REGION Network 2: Orden de marcha desde Panel MC002 - Compresor de Alta ABC3
   RUNG wire#powerrail
      Contact( "PanelCmpAlta".MarchaPanelMC002 )
      I_Contact( "PanelCmpAlta".MantMC002 )
      Coil( "DB-CompAltaDatos".PanMchCmp2 )
   END_RUNG
   // the same network as SCL:
   "DB-CompAltaDatos".PanMchCmp2 := "PanelCmpAlta".MarchaPanelMC002 AND NOT "PanelCmpAlta".MantMC002;
END_REGION

REGION Network 3: Orden de marcha desde Panel MC003 - Compresor de Alta BELLIS
   RUNG wire#powerrail
      Contact( "PanelCmpAlta".MarchaPanelMC003 )
      I_Contact( "PanelCmpAlta".MantMC003 )
      Coil( "DB-CompAltaDatos".PanMchCmp3 )
   END_RUNG
   // the same network as SCL:
   "DB-CompAltaDatos".PanMchCmp3 := "PanelCmpAlta".MarchaPanelMC003 AND NOT "PanelCmpAlta".MantMC003;
END_REGION

REGION Network 4: Orden de marcha desde Panel MC004 - Compresor de Alta ABC4
   RUNG wire#powerrail
      Contact( "PanelCmpAlta".MarchaPanelMC004 )
      I_Contact( "PanelCmpAlta".MantMC004 )
      Coil( "DB-CompAltaDatos".PanMchCmp4 )
   END_RUNG
   // the same network as SCL:
   "DB-CompAltaDatos".PanMchCmp4 := "PanelCmpAlta".MarchaPanelMC004 AND NOT "PanelCmpAlta".MantMC004;
END_REGION

REGION Network 5: Orden de marcha desde Panel MC005 - Compresor de Alta ABC5
   RUNG wire#powerrail
      Contact( "PanelCmpAlta".MarchaPanelMC005 )
      I_Contact( "PanelCmpAlta".MantMC005 )
      Coil( "DB-CompAltaDatos".PanMchCmp5 )
   END_RUNG
   // the same network as SCL:
   "DB-CompAltaDatos".PanMchCmp5 := "PanelCmpAlta".MarchaPanelMC005 AND NOT "PanelCmpAlta".MantMC005;
END_REGION

REGION Network 6: Orden de marcha desde Panel MC005 - Compresor de Alta ABC5
   RUNG wire#powerrail
      Contact( "PanelCmpAlta".MarchaPanelMC006 )
      I_Contact( "PanelCmpAlta".MantMC006 )
      Coil( "DB-CompAltaDatos".PanMchCmp6 )
   END_RUNG
   // the same network as SCL:
   "DB-CompAltaDatos".PanMchCmp6 := "PanelCmpAlta".MarchaPanelMC006 AND NOT "PanelCmpAlta".MantMC006;
END_REGION

REGION Network 7: Salida de mantenimiento compresor 1 / Mantenimiento MC001 - Compresor de Alta ABC2
   RUNG wire#powerrail
      Contact( "PanelCmpAlta".MantMC001 )
      Not()
      Coil( "MC001_MANT" )
   END_RUNG
   // the same network as SCL:
   "MC001_MANT" := NOT "PanelCmpAlta".MantMC001;
END_REGION

REGION Network 8: Salida de mantenimiento compresor 2 / Mantenimiento MC002 - Compresor de Alta ABC3
   RUNG wire#powerrail
      Contact( "PanelCmpAlta".MantMC002 )
      Not()
      Coil( "MC002_MANT" )
   END_RUNG
   // the same network as SCL:
   "MC002_MANT" := NOT "PanelCmpAlta".MantMC002;
END_REGION

REGION Network 9: Salida de mantenimiento compresor 3 / Mantenimiento MC003 - Compresor de Alta BELLIS
   RUNG wire#powerrail
      Contact( "PanelCmpAlta".MantMC003 )
      Not()
      Coil( "MC003_MANT" )
   END_RUNG
   // the same network as SCL:
   "MC003_MANT" := NOT "PanelCmpAlta".MantMC003;
END_REGION

REGION Network 10: Salida de mantenimiento compresor 4 / Mantenimiento MC004 - Compresor de Alta ABC4
   RUNG wire#powerrail
      Contact( "PanelCmpAlta".MantMC004 )
      Not()
      Coil( "MC004_MANT" )
   END_RUNG
   // the same network as SCL:
   "MC004_MANT" := NOT "PanelCmpAlta".MantMC004;
END_REGION

REGION Network 11: Salida de mantenimiento compresor 5 / Mantenimiento MC005 - Compresor de Alta ABC5
   RUNG wire#powerrail
      Contact( "PanelCmpAlta".MantMC005 )
      Not()
      Coil( "MC005_MANT" )
   END_RUNG
   // the same network as SCL:
   "MC005_MANT" := NOT "PanelCmpAlta".MantMC005;
END_REGION

REGION Network 12: Salida de mantenimiento compresor 6 / Mantenimiento MC005 - Compresor de Alta ABC5
   RUNG wire#powerrail
      Contact( "PanelCmpAlta".MantMC006 )
      Not()
      Coil( "MC006_MANT" )
   END_RUNG
   // the same network as SCL:
   "MC006_MANT" := NOT "PanelCmpAlta".MantMC006;
END_REGION

REGION Network 13: Aparentemente obsoleto
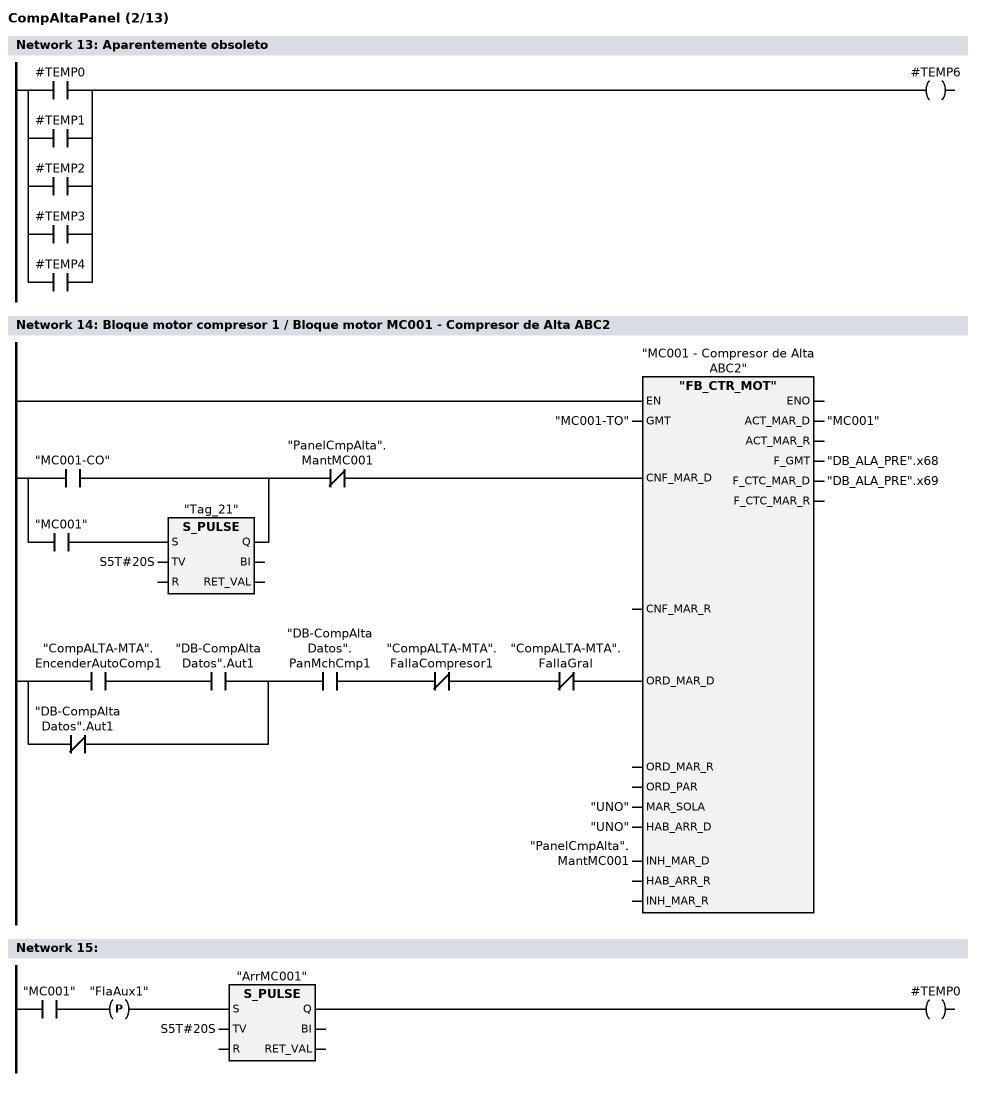
   RUNG wire#powerrail
      Contact( #TEMP0 )
      wire#w1
      Coil( #TEMP6 )
   END_RUNG
   RUNG wire#powerrail
      Contact( #TEMP1 )
   END_RUNG wire#w1
   RUNG wire#powerrail
      Contact( #TEMP2 )
   END_RUNG wire#w1
   RUNG wire#powerrail
      Contact( #TEMP3 )
   END_RUNG wire#w1
   RUNG wire#powerrail
      Contact( #TEMP4 )
   END_RUNG wire#w1
   // the same network as SCL:
   #TEMP6 := #TEMP0 OR #TEMP1 OR #TEMP2 OR #TEMP3 OR #TEMP4;
END_REGION

REGION Network 14: Bloque motor compresor 1 / Bloque motor MC001 - Compresor de Alta ABC2
   RUNG wire#powerrail
      "MC001 - Compresor de Alta ABC2"(CNF_MAR_D := wire#w2, ORD_MAR_D := wire#w4, GMT := "MC001-TO", CNF_MAR_R :=, ORD_MAR_R :=, ORD_PAR :=, MAR_SOLA := "UNO", HAB_ARR_D := "UNO", INH_MAR_D := "PanelCmpAlta".MantMC001, HAB_ARR_R :=, INH_MAR_R :=, ACT_MAR_D => "MC001", ACT_MAR_R =>, F_GMT => "DB_ALA_PRE".x68, F_CTC_MAR_D => "DB_ALA_PRE".x69, F_CTC_MAR_R =>)
   END_RUNG
   RUNG wire#powerrail
      Contact( "MC001-CO" )
      wire#w1
      I_Contact( "PanelCmpAlta".MantMC001 )
   END_RUNG wire#w2
   RUNG wire#powerrail
      Contact( "MC001" )
      S_PULSE(T_NO := "Tag_21", TV := S5T#20S, R :=, BI =>, RET_VAL =>)
   END_RUNG wire#w1
   RUNG wire#powerrail
      Contact( "CompALTA-MTA".EncenderAutoComp1 )
      Contact( "DB-CompAltaDatos".Aut1 )
      wire#w3
      Contact( "DB-CompAltaDatos".PanMchCmp1 )
      I_Contact( "CompALTA-MTA".FallaCompresor1 )
      I_Contact( "CompALTA-MTA".FallaGral )
   END_RUNG wire#w4
   RUNG wire#powerrail
      I_Contact( "DB-CompAltaDatos".Aut1 )
   END_RUNG wire#w3
   // the same network as SCL:
   #_s5time1 := S_PULSE(T_NO := "Tag_21", S := "MC001", TV := S5T#20S, Q => #_w1);
   "MC001 - Compresor de Alta ABC2"(GMT := "MC001-TO",   // "FB_CTR_MOT"
                           CNF_MAR_D := ("MC001-CO" OR #_w1) AND NOT "PanelCmpAlta".MantMC001,
                           ORD_MAR_D := (("CompALTA-MTA".EncenderAutoComp1 AND "DB-CompAltaDatos".Aut1) OR NOT "DB-CompAltaDatos".Aut1) AND "DB-CompAltaDatos".PanMchCmp1 AND NOT "CompALTA-MTA".FallaCompresor1 AND NOT "CompALTA-MTA".FallaGral,
                           MAR_SOLA := "UNO",
                           HAB_ARR_D := "UNO",
                           INH_MAR_D := "PanelCmpAlta".MantMC001,
                           ACT_MAR_D => "MC001",
                           F_GMT => "DB_ALA_PRE".x68,
                           F_CTC_MAR_D => "DB_ALA_PRE".x69);
END_REGION

REGION Network 15
   RUNG wire#powerrail
      Contact( "MC001" )
      P_Trig( "FlaAux1" )
      S_PULSE(T_NO := "ArrMC001", TV := S5T#20S, R :=, BI =>, RET_VAL =>)
      Coil( #TEMP0 )
   END_RUNG
   // the same network as SCL:
   #_w1 := "MC001" AND NOT "FlaAux1";   // rising edge
   "FlaAux1" := "MC001";
   #_s5time1 := S_PULSE(T_NO := "ArrMC001", S := #_w1, TV := S5T#20S, Q => #_w2);
   #TEMP0 := #_w2;
END_REGION

REGION Network 16: Bloque motor compresor 2 / Bloque motor MC002 - Compresor de Alta ABC3
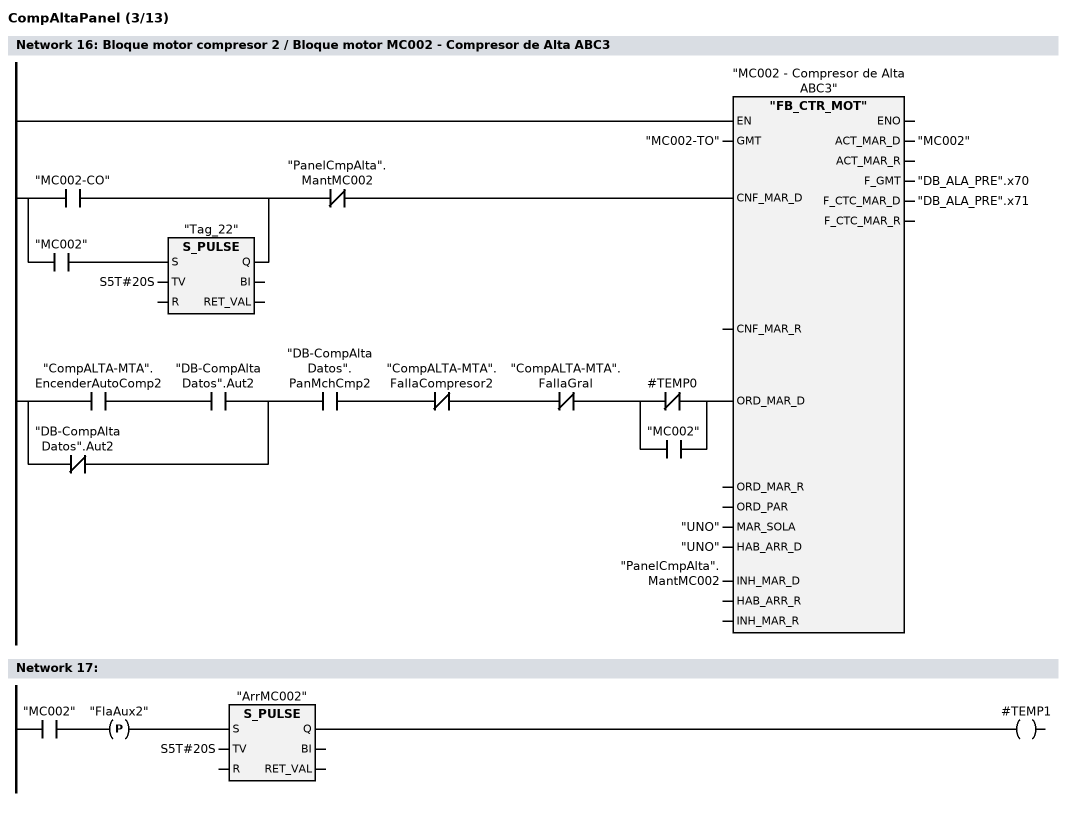
   RUNG wire#powerrail
      "MC002 - Compresor de Alta ABC3"(CNF_MAR_D := wire#w2, ORD_MAR_D := wire#w5, GMT := "MC002-TO", CNF_MAR_R :=, ORD_MAR_R :=, ORD_PAR :=, MAR_SOLA := "UNO", HAB_ARR_D := "UNO", INH_MAR_D := "PanelCmpAlta".MantMC002, HAB_ARR_R :=, INH_MAR_R :=, ACT_MAR_D => "MC002", ACT_MAR_R =>, F_GMT => "DB_ALA_PRE".x70, F_CTC_MAR_D => "DB_ALA_PRE".x71, F_CTC_MAR_R =>)
   END_RUNG
   RUNG wire#powerrail
      Contact( "MC002-CO" )
      wire#w1
      I_Contact( "PanelCmpAlta".MantMC002 )
   END_RUNG wire#w2
   RUNG wire#powerrail
      Contact( "MC002" )
      S_PULSE(T_NO := "Tag_22", TV := S5T#20S, R :=, BI =>, RET_VAL =>)
   END_RUNG wire#w1
   RUNG wire#powerrail
      Contact( "CompALTA-MTA".EncenderAutoComp2 )
      Contact( "DB-CompAltaDatos".Aut2 )
      wire#w3
      Contact( "DB-CompAltaDatos".PanMchCmp2 )
      I_Contact( "CompALTA-MTA".FallaCompresor2 )
      I_Contact( "CompALTA-MTA".FallaGral )
      wire#w4
      I_Contact( #TEMP0 )
   END_RUNG wire#w5
   RUNG wire#powerrail
      I_Contact( "DB-CompAltaDatos".Aut2 )
   END_RUNG wire#w3
   RUNG wire#w4
      Contact( "MC002" )
   END_RUNG wire#w5
   // the same network as SCL:
   #_s5time1 := S_PULSE(T_NO := "Tag_22", S := "MC002", TV := S5T#20S, Q => #_w1);
   "MC002 - Compresor de Alta ABC3"(GMT := "MC002-TO",   // "FB_CTR_MOT"
                           CNF_MAR_D := ("MC002-CO" OR #_w1) AND NOT "PanelCmpAlta".MantMC002,
                           ORD_MAR_D := (("CompALTA-MTA".EncenderAutoComp2 AND "DB-CompAltaDatos".Aut2) OR NOT "DB-CompAltaDatos".Aut2) AND "DB-CompAltaDatos".PanMchCmp2 AND NOT "CompALTA-MTA".FallaCompresor2 AND NOT "CompALTA-MTA".FallaGral AND (NOT #TEMP0 OR "MC002"),
                           MAR_SOLA := "UNO",
                           HAB_ARR_D := "UNO",
                           INH_MAR_D := "PanelCmpAlta".MantMC002,
                           ACT_MAR_D => "MC002",
                           F_GMT => "DB_ALA_PRE".x70,
                           F_CTC_MAR_D => "DB_ALA_PRE".x71);
END_REGION

REGION Network 17
   RUNG wire#powerrail
      Contact( "MC002" )
      P_Trig( "FlaAux2" )
      S_PULSE(T_NO := "ArrMC002", TV := S5T#20S, R :=, BI =>, RET_VAL =>)
      Coil( #TEMP1 )
   END_RUNG
   // the same network as SCL:
   #_w1 := "MC002" AND NOT "FlaAux2";   // rising edge
   "FlaAux2" := "MC002";
   #_s5time1 := S_PULSE(T_NO := "ArrMC002", S := #_w1, TV := S5T#20S, Q => #_w2);
   #TEMP1 := #_w2;
END_REGION

REGION Network 18: Bloque motor compresor 3 / Bloque motor MC003 - Compresor de Alta BELLIS
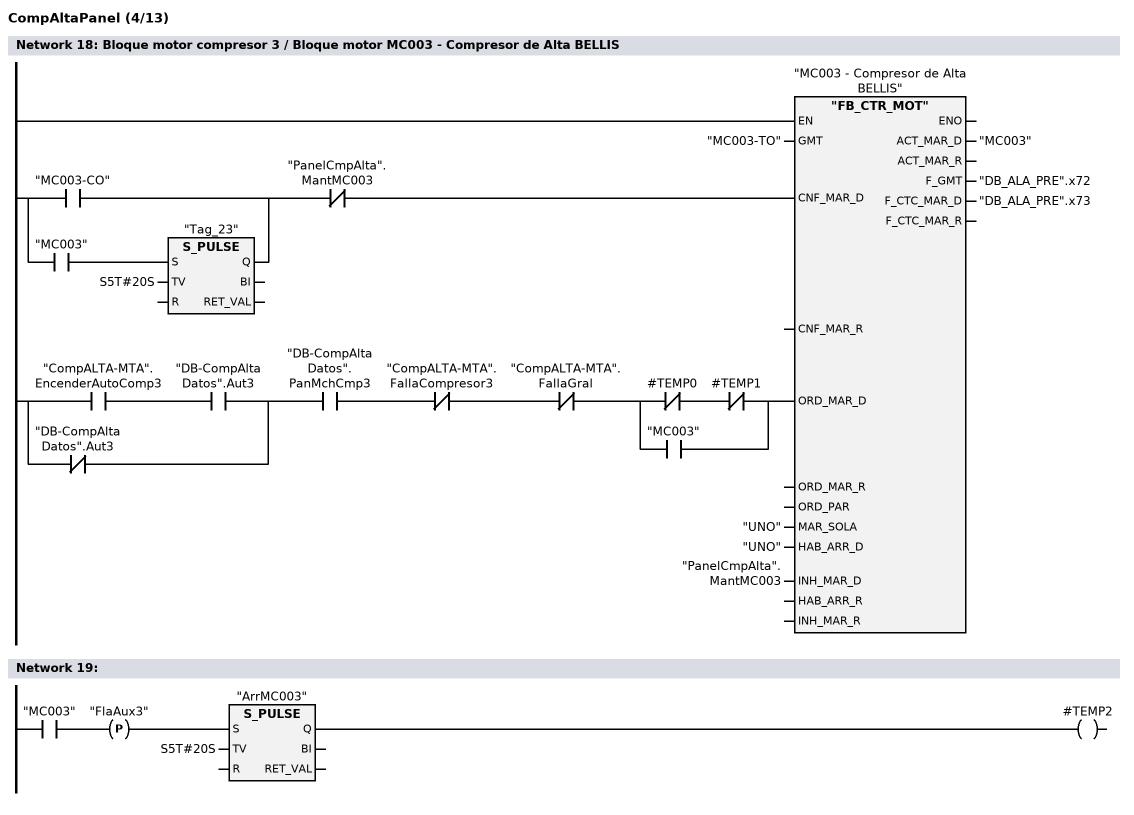
   RUNG wire#powerrail
      "MC003 - Compresor de Alta BELLIS"(CNF_MAR_D := wire#w2, ORD_MAR_D := wire#w5, GMT := "MC003-TO", CNF_MAR_R :=, ORD_MAR_R :=, ORD_PAR :=, MAR_SOLA := "UNO", HAB_ARR_D := "UNO", INH_MAR_D := "PanelCmpAlta".MantMC003, HAB_ARR_R :=, INH_MAR_R :=, ACT_MAR_D => "MC003", ACT_MAR_R =>, F_GMT => "DB_ALA_PRE".x72, F_CTC_MAR_D => "DB_ALA_PRE".x73, F_CTC_MAR_R =>)
   END_RUNG
   RUNG wire#powerrail
      Contact( "MC003-CO" )
      wire#w1
      I_Contact( "PanelCmpAlta".MantMC003 )
   END_RUNG wire#w2
   RUNG wire#powerrail
      Contact( "MC003" )
      S_PULSE(T_NO := "Tag_23", TV := S5T#20S, R :=, BI =>, RET_VAL =>)
   END_RUNG wire#w1
   RUNG wire#powerrail
      Contact( "CompALTA-MTA".EncenderAutoComp3 )
      Contact( "DB-CompAltaDatos".Aut3 )
      wire#w3
      Contact( "DB-CompAltaDatos".PanMchCmp3 )
      I_Contact( "CompALTA-MTA".FallaCompresor3 )
      I_Contact( "CompALTA-MTA".FallaGral )
      wire#w4
      I_Contact( #TEMP0 )
      I_Contact( #TEMP1 )
   END_RUNG wire#w5
   RUNG wire#powerrail
      I_Contact( "DB-CompAltaDatos".Aut3 )
   END_RUNG wire#w3
   RUNG wire#w4
      Contact( "MC003" )
   END_RUNG wire#w5
   // the same network as SCL:
   #_s5time1 := S_PULSE(T_NO := "Tag_23", S := "MC003", TV := S5T#20S, Q => #_w1);
   "MC003 - Compresor de Alta BELLIS"(GMT := "MC003-TO",   // "FB_CTR_MOT"
                           CNF_MAR_D := ("MC003-CO" OR #_w1) AND NOT "PanelCmpAlta".MantMC003,
                           ORD_MAR_D := (("CompALTA-MTA".EncenderAutoComp3 AND "DB-CompAltaDatos".Aut3) OR NOT "DB-CompAltaDatos".Aut3) AND "DB-CompAltaDatos".PanMchCmp3 AND NOT "CompALTA-MTA".FallaCompresor3 AND NOT "CompALTA-MTA".FallaGral AND ((NOT #TEMP0 AND NOT #TEMP1) OR "MC003"),
                           MAR_SOLA := "UNO",
                           HAB_ARR_D := "UNO",
                           INH_MAR_D := "PanelCmpAlta".MantMC003,
                           ACT_MAR_D => "MC003",
                           F_GMT => "DB_ALA_PRE".x72,
                           F_CTC_MAR_D => "DB_ALA_PRE".x73);
END_REGION

REGION Network 19
   RUNG wire#powerrail
      Contact( "MC003" )
      P_Trig( "FlaAux3" )
      S_PULSE(T_NO := "ArrMC003", TV := S5T#20S, R :=, BI =>, RET_VAL =>)
      Coil( #TEMP2 )
   END_RUNG
   // the same network as SCL:
   #_w1 := "MC003" AND NOT "FlaAux3";   // rising edge
   "FlaAux3" := "MC003";
   #_s5time1 := S_PULSE(T_NO := "ArrMC003", S := #_w1, TV := S5T#20S, Q => #_w2);
   #TEMP2 := #_w2;
END_REGION

REGION Network 20: Bloque motor compresor 4 / Bloque motor MC004 - Compresor de Alta ABC4
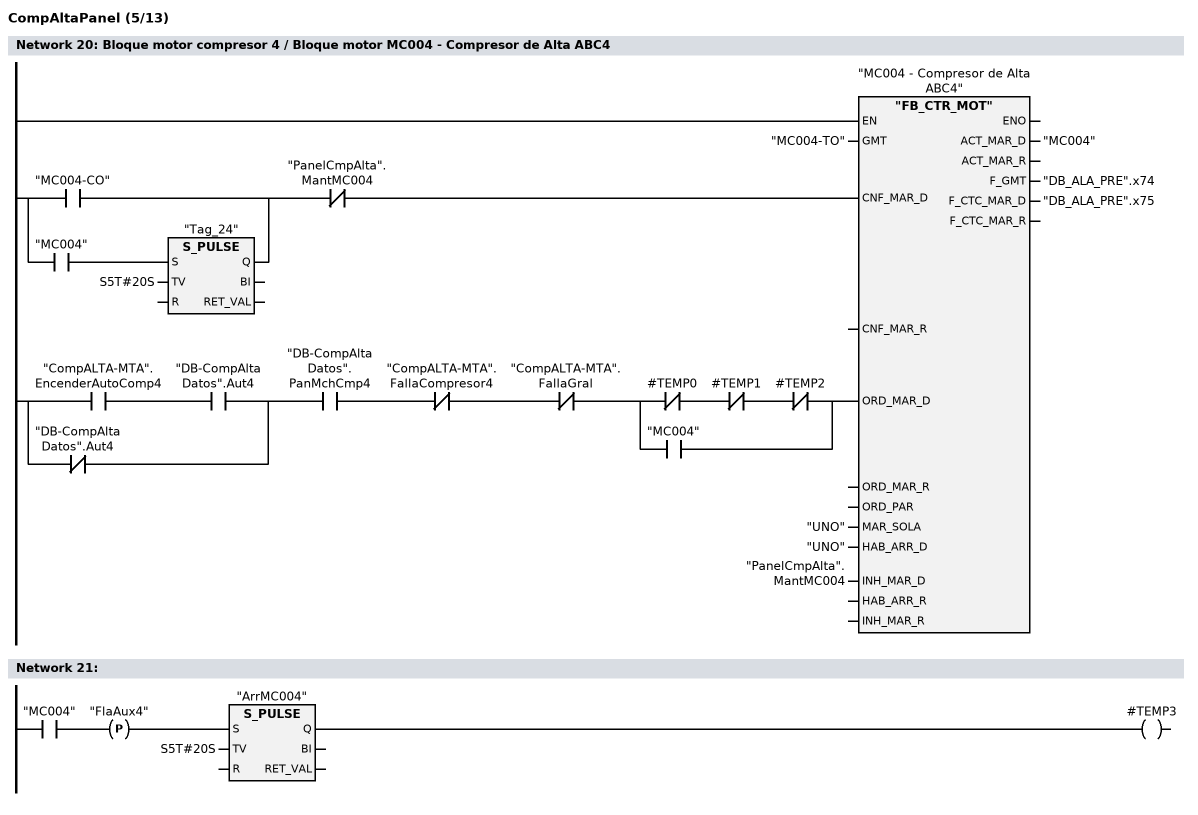
   RUNG wire#powerrail
      "MC004 - Compresor de Alta ABC4"(CNF_MAR_D := wire#w2, ORD_MAR_D := wire#w5, GMT := "MC004-TO", CNF_MAR_R :=, ORD_MAR_R :=, ORD_PAR :=, MAR_SOLA := "UNO", HAB_ARR_D := "UNO", INH_MAR_D := "PanelCmpAlta".MantMC004, HAB_ARR_R :=, INH_MAR_R :=, ACT_MAR_D => "MC004", ACT_MAR_R =>, F_GMT => "DB_ALA_PRE".x74, F_CTC_MAR_D => "DB_ALA_PRE".x75, F_CTC_MAR_R =>)
   END_RUNG
   RUNG wire#powerrail
      Contact( "MC004-CO" )
      wire#w1
      I_Contact( "PanelCmpAlta".MantMC004 )
   END_RUNG wire#w2
   RUNG wire#powerrail
      Contact( "MC004" )
      S_PULSE(T_NO := "Tag_24", TV := S5T#20S, R :=, BI =>, RET_VAL =>)
   END_RUNG wire#w1
   RUNG wire#powerrail
      Contact( "CompALTA-MTA".EncenderAutoComp4 )
      Contact( "DB-CompAltaDatos".Aut4 )
      wire#w3
      Contact( "DB-CompAltaDatos".PanMchCmp4 )
      I_Contact( "CompALTA-MTA".FallaCompresor4 )
      I_Contact( "CompALTA-MTA".FallaGral )
      wire#w4
      I_Contact( #TEMP0 )
      I_Contact( #TEMP1 )
      I_Contact( #TEMP2 )
   END_RUNG wire#w5
   RUNG wire#powerrail
      I_Contact( "DB-CompAltaDatos".Aut4 )
   END_RUNG wire#w3
   RUNG wire#w4
      Contact( "MC004" )
   END_RUNG wire#w5
   // the same network as SCL:
   #_s5time1 := S_PULSE(T_NO := "Tag_24", S := "MC004", TV := S5T#20S, Q => #_w1);
   "MC004 - Compresor de Alta ABC4"(GMT := "MC004-TO",   // "FB_CTR_MOT"
                           CNF_MAR_D := ("MC004-CO" OR #_w1) AND NOT "PanelCmpAlta".MantMC004,
                           ORD_MAR_D := (("CompALTA-MTA".EncenderAutoComp4 AND "DB-CompAltaDatos".Aut4) OR NOT "DB-CompAltaDatos".Aut4) AND "DB-CompAltaDatos".PanMchCmp4 AND NOT "CompALTA-MTA".FallaCompresor4 AND NOT "CompALTA-MTA".FallaGral AND ((NOT #TEMP0 AND NOT #TEMP1 AND NOT #TEMP2) OR "MC004"),
                           MAR_SOLA := "UNO",
                           HAB_ARR_D := "UNO",
                           INH_MAR_D := "PanelCmpAlta".MantMC004,
                           ACT_MAR_D => "MC004",
                           F_GMT => "DB_ALA_PRE".x74,
                           F_CTC_MAR_D => "DB_ALA_PRE".x75);
END_REGION

REGION Network 21
   RUNG wire#powerrail
      Contact( "MC004" )
      P_Trig( "FlaAux4" )
      S_PULSE(T_NO := "ArrMC004", TV := S5T#20S, R :=, BI =>, RET_VAL =>)
      Coil( #TEMP3 )
   END_RUNG
   // the same network as SCL:
   #_w1 := "MC004" AND NOT "FlaAux4";   // rising edge
   "FlaAux4" := "MC004";
   #_s5time1 := S_PULSE(T_NO := "ArrMC004", S := #_w1, TV := S5T#20S, Q => #_w2);
   #TEMP3 := #_w2;
END_REGION

REGION Network 22: Bloque motor compresor 5 / Bloque motor MC005 - Compresor de Alta ABC5
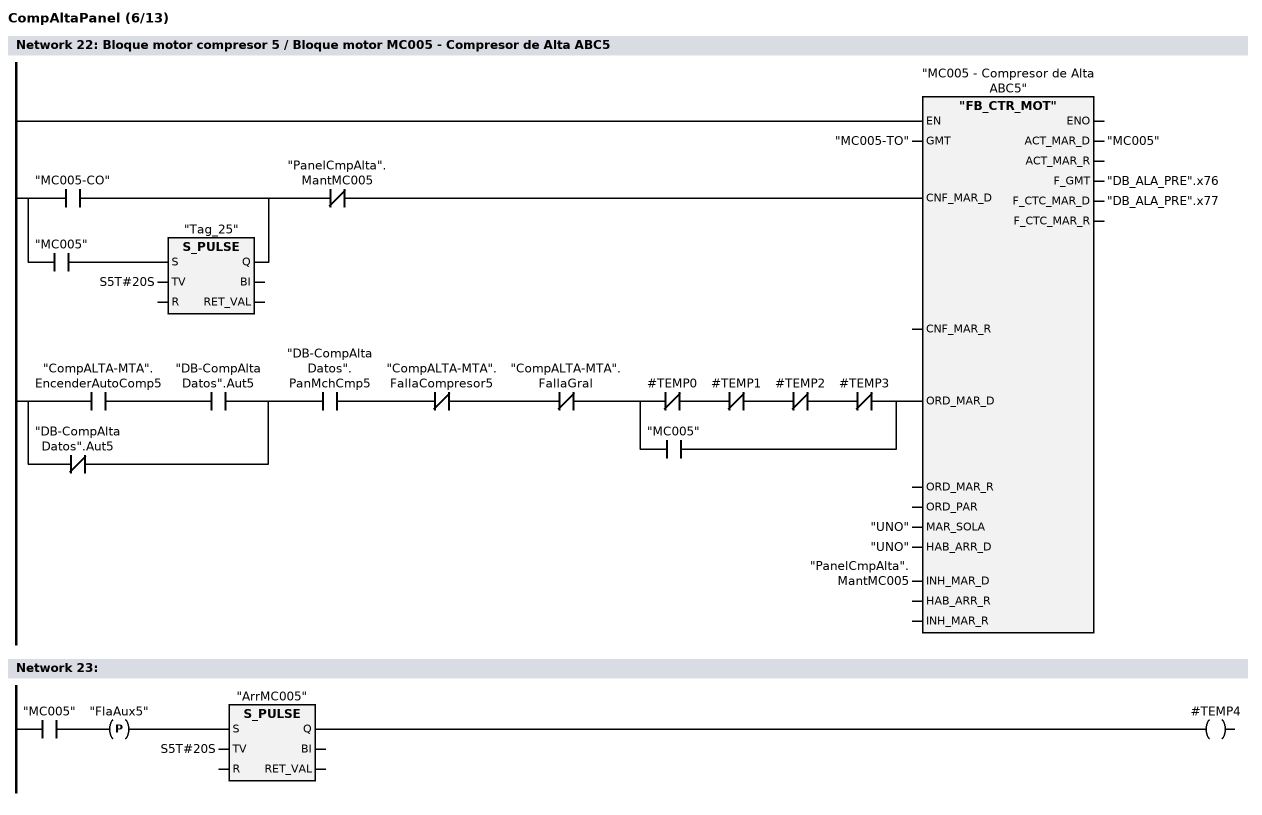
   RUNG wire#powerrail
      "MC005 - Compresor de Alta ABC5"(CNF_MAR_D := wire#w2, ORD_MAR_D := wire#w5, GMT := "MC005-TO", CNF_MAR_R :=, ORD_MAR_R :=, ORD_PAR :=, MAR_SOLA := "UNO", HAB_ARR_D := "UNO", INH_MAR_D := "PanelCmpAlta".MantMC005, HAB_ARR_R :=, INH_MAR_R :=, ACT_MAR_D => "MC005", ACT_MAR_R =>, F_GMT => "DB_ALA_PRE".x76, F_CTC_MAR_D => "DB_ALA_PRE".x77, F_CTC_MAR_R =>)
   END_RUNG
   RUNG wire#powerrail
      Contact( "MC005-CO" )
      wire#w1
      I_Contact( "PanelCmpAlta".MantMC005 )
   END_RUNG wire#w2
   RUNG wire#powerrail
      Contact( "MC005" )
      S_PULSE(T_NO := "Tag_25", TV := S5T#20S, R :=, BI =>, RET_VAL =>)
   END_RUNG wire#w1
   RUNG wire#powerrail
      Contact( "CompALTA-MTA".EncenderAutoComp5 )
      Contact( "DB-CompAltaDatos".Aut5 )
      wire#w3
      Contact( "DB-CompAltaDatos".PanMchCmp5 )
      I_Contact( "CompALTA-MTA".FallaCompresor5 )
      I_Contact( "CompALTA-MTA".FallaGral )
      wire#w4
      I_Contact( #TEMP0 )
      I_Contact( #TEMP1 )
      I_Contact( #TEMP2 )
      I_Contact( #TEMP3 )
   END_RUNG wire#w5
   RUNG wire#powerrail
      I_Contact( "DB-CompAltaDatos".Aut5 )
   END_RUNG wire#w3
   RUNG wire#w4
      Contact( "MC005" )
   END_RUNG wire#w5
   // the same network as SCL:
   #_s5time1 := S_PULSE(T_NO := "Tag_25", S := "MC005", TV := S5T#20S, Q => #_w1);
   "MC005 - Compresor de Alta ABC5"(GMT := "MC005-TO",   // "FB_CTR_MOT"
                           CNF_MAR_D := ("MC005-CO" OR #_w1) AND NOT "PanelCmpAlta".MantMC005,
                           ORD_MAR_D := (("CompALTA-MTA".EncenderAutoComp5 AND "DB-CompAltaDatos".Aut5) OR NOT "DB-CompAltaDatos".Aut5) AND "DB-CompAltaDatos".PanMchCmp5 AND NOT "CompALTA-MTA".FallaCompresor5 AND NOT "CompALTA-MTA".FallaGral AND ((NOT #TEMP0 AND NOT #TEMP1 AND NOT #TEMP2 AND NOT #TEMP3) OR "MC005"),
                           MAR_SOLA := "UNO",
                           HAB_ARR_D := "UNO",
                           INH_MAR_D := "PanelCmpAlta".MantMC005,
                           ACT_MAR_D => "MC005",
                           F_GMT => "DB_ALA_PRE".x76,
                           F_CTC_MAR_D => "DB_ALA_PRE".x77);
END_REGION

REGION Network 23
   RUNG wire#powerrail
      Contact( "MC005" )
      P_Trig( "FlaAux5" )
      S_PULSE(T_NO := "ArrMC005", TV := S5T#20S, R :=, BI =>, RET_VAL =>)
      Coil( #TEMP4 )
   END_RUNG
   // the same network as SCL:
   #_w1 := "MC005" AND NOT "FlaAux5";   // rising edge
   "FlaAux5" := "MC005";
   #_s5time1 := S_PULSE(T_NO := "ArrMC005", S := #_w1, TV := S5T#20S, Q => #_w2);
   #TEMP4 := #_w2;
END_REGION

REGION Network 24: Bloque motor compresor 6 / Bloque motor MC005 - Compresor de Alta ABC5
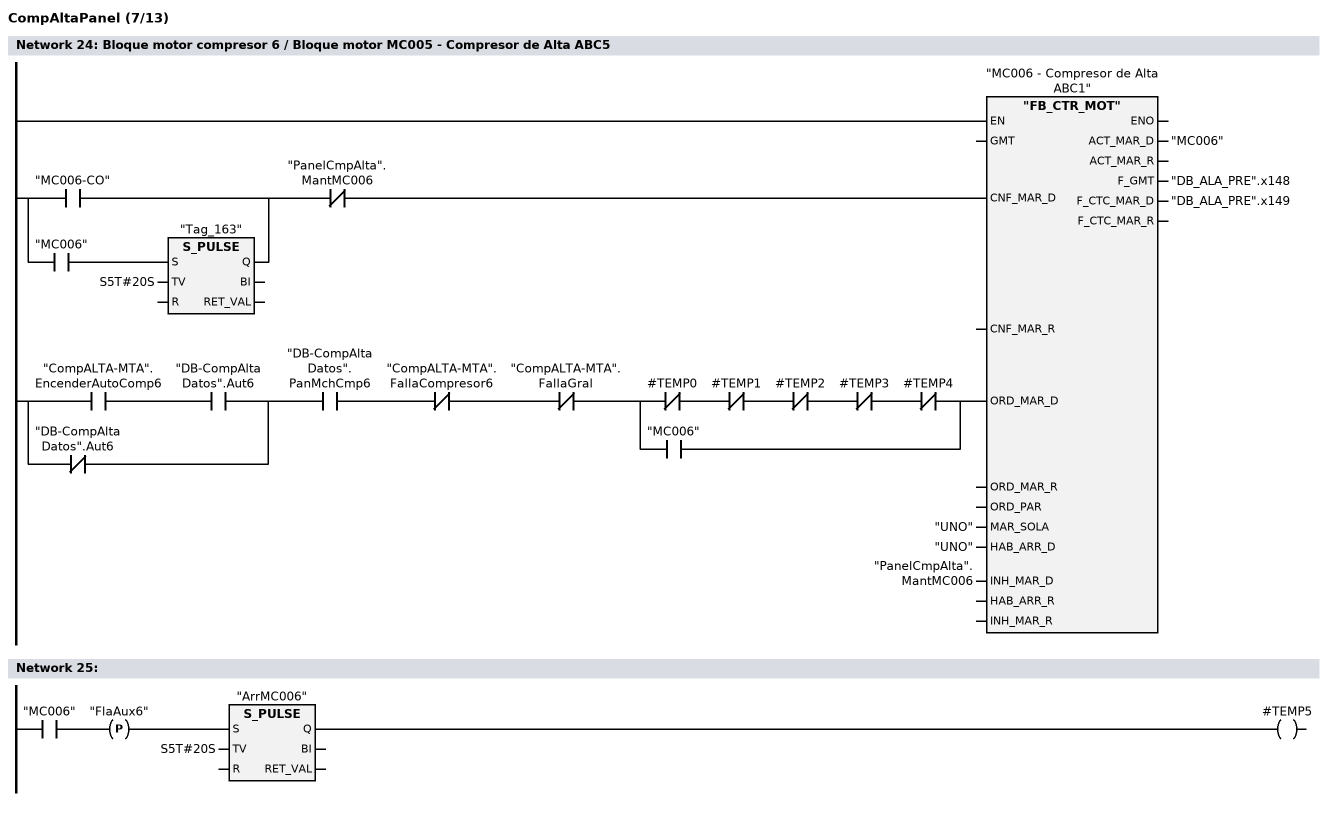
   RUNG wire#powerrail
      "MC006 - Compresor de Alta ABC1"(CNF_MAR_D := wire#w2, ORD_MAR_D := wire#w5, GMT :=, CNF_MAR_R :=, ORD_MAR_R :=, ORD_PAR :=, MAR_SOLA := "UNO", HAB_ARR_D := "UNO", INH_MAR_D := "PanelCmpAlta".MantMC006, HAB_ARR_R :=, INH_MAR_R :=, ACT_MAR_D => "MC006", ACT_MAR_R =>, F_GMT => "DB_ALA_PRE".x148, F_CTC_MAR_D => "DB_ALA_PRE".x149, F_CTC_MAR_R =>)
   END_RUNG
   RUNG wire#powerrail
      Contact( "MC006-CO" )
      wire#w1
      I_Contact( "PanelCmpAlta".MantMC006 )
   END_RUNG wire#w2
   RUNG wire#powerrail
      Contact( "MC006" )
      S_PULSE(T_NO := "Tag_163", TV := S5T#20S, R :=, BI =>, RET_VAL =>)
   END_RUNG wire#w1
   RUNG wire#powerrail
      Contact( "CompALTA-MTA".EncenderAutoComp6 )
      Contact( "DB-CompAltaDatos".Aut6 )
      wire#w3
      Contact( "DB-CompAltaDatos".PanMchCmp6 )
      I_Contact( "CompALTA-MTA".FallaCompresor6 )
      I_Contact( "CompALTA-MTA".FallaGral )
      wire#w4
      I_Contact( #TEMP0 )
      I_Contact( #TEMP1 )
      I_Contact( #TEMP2 )
      I_Contact( #TEMP3 )
      I_Contact( #TEMP4 )
   END_RUNG wire#w5
   RUNG wire#powerrail
      I_Contact( "DB-CompAltaDatos".Aut6 )
   END_RUNG wire#w3
   RUNG wire#w4
      Contact( "MC006" )
   END_RUNG wire#w5
   // the same network as SCL:
   #_s5time1 := S_PULSE(T_NO := "Tag_163", S := "MC006", TV := S5T#20S, Q => #_w1);
   "MC006 - Compresor de Alta ABC1"(CNF_MAR_D := ("MC006-CO" OR #_w1) AND NOT "PanelCmpAlta".MantMC006,   // "FB_CTR_MOT"
                           ORD_MAR_D := (("CompALTA-MTA".EncenderAutoComp6 AND "DB-CompAltaDatos".Aut6) OR NOT "DB-CompAltaDatos".Aut6) AND "DB-CompAltaDatos".PanMchCmp6 AND NOT "CompALTA-MTA".FallaCompresor6 AND NOT "CompALTA-MTA".FallaGral AND ((NOT #TEMP0 AND NOT #TEMP1 AND NOT #TEMP2 AND NOT #TEMP3 AND NOT #TEMP4) OR "MC006"),
                           MAR_SOLA := "UNO",
                           HAB_ARR_D := "UNO",
                           INH_MAR_D := "PanelCmpAlta".MantMC006,
                           ACT_MAR_D => "MC006",
                           F_GMT => "DB_ALA_PRE".x148,
                           F_CTC_MAR_D => "DB_ALA_PRE".x149);
END_REGION

REGION Network 25
   RUNG wire#powerrail
      Contact( "MC006" )
      P_Trig( "FlaAux6" )
      S_PULSE(T_NO := "ArrMC006", TV := S5T#20S, R :=, BI =>, RET_VAL =>)
      Coil( #TEMP5 )
   END_RUNG
   // the same network as SCL:
   #_w1 := "MC006" AND NOT "FlaAux6";   // rising edge
   "FlaAux6" := "MC006";
   #_s5time1 := S_PULSE(T_NO := "ArrMC006", S := #_w1, TV := S5T#20S, Q => #_w2);
   #TEMP5 := #_w2;
END_REGION

REGION Network 26: Bloque de animación motor compresor 1 / Animación Motor MC001 - Compresor de Alta ABC2
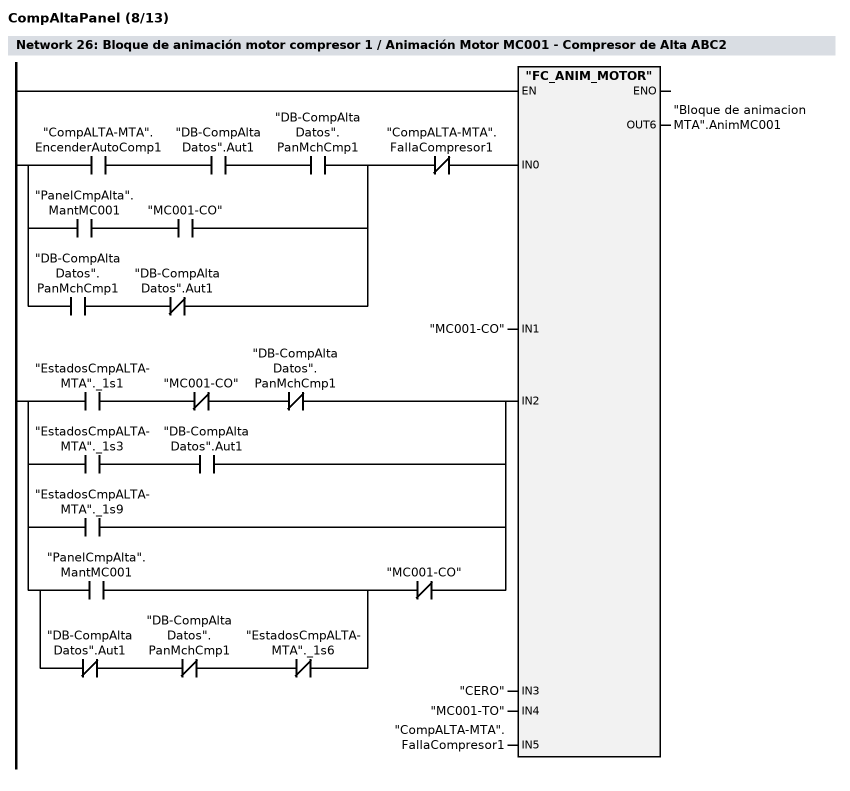
   RUNG wire#powerrail
      "FC_ANIM_MOTOR"(IN0 := wire#w2, IN2 := wire#w4, IN1 := "MC001-CO", IN3 := "CERO", IN4 := "MC001-TO", IN5 := "CompALTA-MTA".FallaCompresor1, OUT6 => "Bloque de animacion MTA".AnimMC001)
   END_RUNG
   RUNG wire#powerrail
      Contact( "CompALTA-MTA".EncenderAutoComp1 )
      Contact( "DB-CompAltaDatos".Aut1 )
      Contact( "DB-CompAltaDatos".PanMchCmp1 )
      wire#w1
      I_Contact( "CompALTA-MTA".FallaCompresor1 )
   END_RUNG wire#w2
   RUNG wire#powerrail
      Contact( "PanelCmpAlta".MantMC001 )
      Contact( "MC001-CO" )
   END_RUNG wire#w1
   RUNG wire#powerrail
      Contact( "DB-CompAltaDatos".PanMchCmp1 )
      I_Contact( "DB-CompAltaDatos".Aut1 )
   END_RUNG wire#w1
   RUNG wire#powerrail
      Contact( "EstadosCmpALTA-MTA"._1s1 )
      I_Contact( "MC001-CO" )
      I_Contact( "DB-CompAltaDatos".PanMchCmp1 )
   END_RUNG wire#w4
   RUNG wire#powerrail
      Contact( "EstadosCmpALTA-MTA"._1s3 )
      Contact( "DB-CompAltaDatos".Aut1 )
   END_RUNG wire#w4
   RUNG wire#powerrail
      Contact( "EstadosCmpALTA-MTA"._1s9 )
   END_RUNG wire#w4
   RUNG wire#powerrail
      Contact( "PanelCmpAlta".MantMC001 )
      wire#w3
      I_Contact( "MC001-CO" )
   END_RUNG wire#w4
   RUNG wire#powerrail
      I_Contact( "DB-CompAltaDatos".Aut1 )
      I_Contact( "DB-CompAltaDatos".PanMchCmp1 )
      I_Contact( "EstadosCmpALTA-MTA"._1s6 )
   END_RUNG wire#w3
   // the same network as SCL:
   "FC_ANIM_MOTOR"(IN0 := (("CompALTA-MTA".EncenderAutoComp1 AND "DB-CompAltaDatos".Aut1 AND "DB-CompAltaDatos".PanMchCmp1) OR ("PanelCmpAlta".MantMC001 AND "MC001-CO") OR ("DB-CompAltaDatos".PanMchCmp1 AND NOT "DB-CompAltaDatos".Aut1)) AND NOT "CompALTA-MTA".FallaCompresor1,
                   IN1 := "MC001-CO",
                   IN2 := ("EstadosCmpALTA-MTA"._1s1 AND NOT "MC001-CO" AND NOT "DB-CompAltaDatos".PanMchCmp1) OR ("EstadosCmpALTA-MTA"._1s3 AND "DB-CompAltaDatos".Aut1) OR "EstadosCmpALTA-MTA"._1s9 OR (("PanelCmpAlta".MantMC001 OR (NOT "DB-CompAltaDatos".Aut1 AND NOT "DB-CompAltaDatos".PanMchCmp1 AND NOT "EstadosCmpALTA-MTA"._1s6)) AND NOT "MC001-CO"),
                   IN3 := "CERO",
                   IN4 := "MC001-TO",
                   IN5 := "CompALTA-MTA".FallaCompresor1,
                   OUT6 => "Bloque de animacion MTA".AnimMC001);
END_REGION

REGION Network 27: Bloque de animación motor compresor 2 / Animación Motor MC002 - Compresor de Alta ABC3
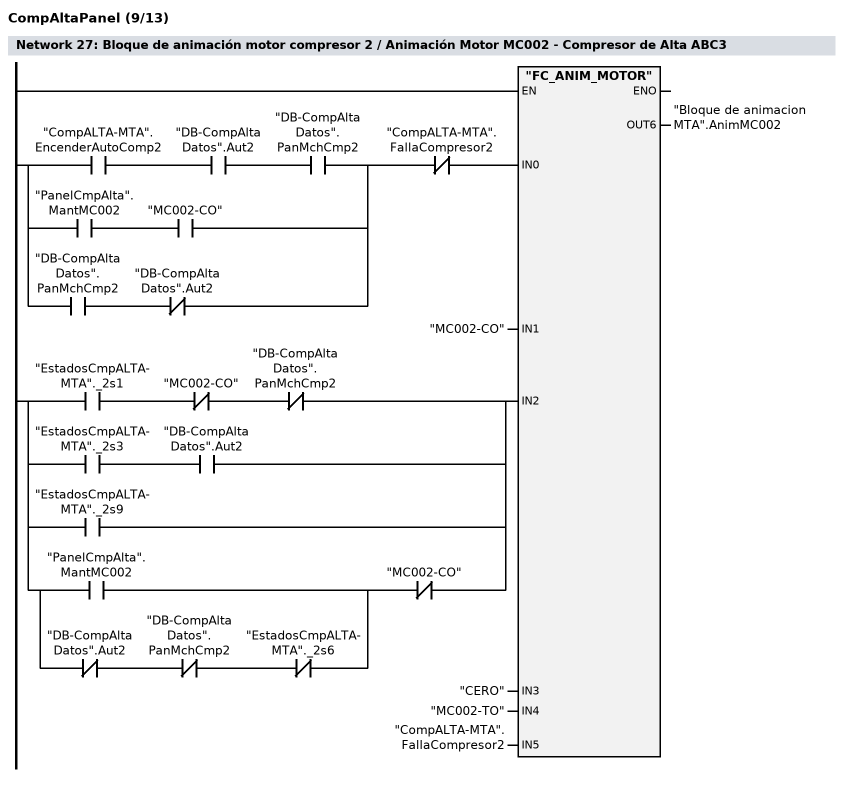
   RUNG wire#powerrail
      "FC_ANIM_MOTOR"(IN0 := wire#w2, IN2 := wire#w4, IN1 := "MC002-CO", IN3 := "CERO", IN4 := "MC002-TO", IN5 := "CompALTA-MTA".FallaCompresor2, OUT6 => "Bloque de animacion MTA".AnimMC002)
   END_RUNG
   RUNG wire#powerrail
      Contact( "CompALTA-MTA".EncenderAutoComp2 )
      Contact( "DB-CompAltaDatos".Aut2 )
      Contact( "DB-CompAltaDatos".PanMchCmp2 )
      wire#w1
      I_Contact( "CompALTA-MTA".FallaCompresor2 )
   END_RUNG wire#w2
   RUNG wire#powerrail
      Contact( "PanelCmpAlta".MantMC002 )
      Contact( "MC002-CO" )
   END_RUNG wire#w1
   RUNG wire#powerrail
      Contact( "DB-CompAltaDatos".PanMchCmp2 )
      I_Contact( "DB-CompAltaDatos".Aut2 )
   END_RUNG wire#w1
   RUNG wire#powerrail
      Contact( "EstadosCmpALTA-MTA"._2s1 )
      I_Contact( "MC002-CO" )
      I_Contact( "DB-CompAltaDatos".PanMchCmp2 )
   END_RUNG wire#w4
   RUNG wire#powerrail
      Contact( "EstadosCmpALTA-MTA"._2s3 )
      Contact( "DB-CompAltaDatos".Aut2 )
   END_RUNG wire#w4
   RUNG wire#powerrail
      Contact( "EstadosCmpALTA-MTA"._2s9 )
   END_RUNG wire#w4
   RUNG wire#powerrail
      Contact( "PanelCmpAlta".MantMC002 )
      wire#w3
      I_Contact( "MC002-CO" )
   END_RUNG wire#w4
   RUNG wire#powerrail
      I_Contact( "DB-CompAltaDatos".Aut2 )
      I_Contact( "DB-CompAltaDatos".PanMchCmp2 )
      I_Contact( "EstadosCmpALTA-MTA"._2s6 )
   END_RUNG wire#w3
   // the same network as SCL:
   "FC_ANIM_MOTOR"(IN0 := (("CompALTA-MTA".EncenderAutoComp2 AND "DB-CompAltaDatos".Aut2 AND "DB-CompAltaDatos".PanMchCmp2) OR ("PanelCmpAlta".MantMC002 AND "MC002-CO") OR ("DB-CompAltaDatos".PanMchCmp2 AND NOT "DB-CompAltaDatos".Aut2)) AND NOT "CompALTA-MTA".FallaCompresor2,
                   IN1 := "MC002-CO",
                   IN2 := ("EstadosCmpALTA-MTA"._2s1 AND NOT "MC002-CO" AND NOT "DB-CompAltaDatos".PanMchCmp2) OR ("EstadosCmpALTA-MTA"._2s3 AND "DB-CompAltaDatos".Aut2) OR "EstadosCmpALTA-MTA"._2s9 OR (("PanelCmpAlta".MantMC002 OR (NOT "DB-CompAltaDatos".Aut2 AND NOT "DB-CompAltaDatos".PanMchCmp2 AND NOT "EstadosCmpALTA-MTA"._2s6)) AND NOT "MC002-CO"),
                   IN3 := "CERO",
                   IN4 := "MC002-TO",
                   IN5 := "CompALTA-MTA".FallaCompresor2,
                   OUT6 => "Bloque de animacion MTA".AnimMC002);
END_REGION

REGION Network 28: Bloque de animación motor compresor 3 / Animación Motor MC003 - Compresor de Alta BELLIS
